   2137: '600-TX-433 APT O2 MONITOR - LOW LOW', class Tank Control Warnings, trigger "2062_Warning_Data_BTCS_WARNING_WORD_01" bit 9
   2138: 'TIT-436 2 PORT BWT TEMP - HIGH', class Tank Control Warnings, trigger "2062_Warning_Data_BTCS_WARNING_WORD_01" bit 10
   2139: 'TIT-436 2 STARBOARD BWT TEMP - HIGH', class Tank Control Warnings, trigger "2062_Warning_Data_BTCS_WARNING_WORD_01" bit 11
   2140: 'BTCS_WARNING_WORD_01_BIT_4', class Tank Control Warnings, trigger "2062_Warning_Data_BTCS_WARNING_WORD_01" bit 12
   2141: 'BTCS_WARNING_WORD_01_BIT_5', class Tank Control Warnings, trigger "2062_Warning_Data_BTCS_WARNING_WORD_01" bit 13
   2142: 'BTCS_WARNING_WORD_01_BIT_6', class Tank Control Warnings, trigger "2062_Warning_Data_BTCS_WARNING_WORD_01" bit 14
   2143: 'BTCS_WARNING_WORD_01_BIT_7', class Tank Control Warnings, trigger "2062_Warning_Data_BTCS_WARNING_WORD_01" bit 15
   2144: 'TT-426 1 FOR PEACK TANK TEMPERATURE - HIGH', class Tank Control Warnings, trigger "2062_Warning_Data_BTCS_WARNING_WORD_02" bit 0
   2145: 'TT-426 1 PORT TANK TEMPERATURE - HIGH', class Tank Control Warnings, trigger "2062_Warning_Data_BTCS_WARNING_WORD_02" bit 1
   2146: 'TT-426 1 STARBOARD TANK TEMPERATURE - HIGH', class Tank Control Warnings, trigger "2062_Warning_Data_BTCS_WARNING_WORD_02" bit 2
   2147: 'TT-426 3 PORT TANK TEMPERATURE - HIGH', class Tank Control Warnings, trigger "2062_Warning_Data_BTCS_WARNING_WORD_02" bit 3
   2148: 'TT-426 3 STARBOARD TANK TEMPERATURE - HIGH', class Tank Control Warnings, trigger "2062_Warning_Data_BTCS_WARNING_WORD_02" bit 4
   2149: 'TT-426 4 PORT TANK TEMPERATURE - HIGH', class Tank Control Warnings, trigger "2062_Warning_Data_BTCS_WARNING_WORD_02" bit 5
   2150: 'TT-426 4 STARBOARD TANK TEMPERATURE - HIGH', class Tank Control Warnings, trigger "2062_Warning_Data_BTCS_WARNING_WORD_02" bit 6
   2151: 'TT-426 5 PORT TANK TEMPERATURE - HIGH', class Tank Control Warnings, trigger "2062_Warning_Data_BTCS_WARNING_WORD_02" bit 7
   2152: 'PIT-415 2 PORT DECK IG PRESSURE - LOW', class Tank Control Warnings, trigger "2062_Warning_Data_BTCS_WARNING_WORD_02" bit 8
   2153: 'PIT-415 2 PORT DECK IG PRESSURE - HIGH', class Tank Control Warnings, trigger "2062_Warning_Data_BTCS_WARNING_WORD_02" bit 9
   2154: 'PIT-415 2 STARBOARD DECK IG PRESSURE - LOW', class Tank Control Warnings, trigger "2062_Warning_Data_BTCS_WARNING_WORD_02" bit 10
   2155: 'PIT-415 STARBOARD DECK IG PRESSURE - HIGH', class Tank Control Warnings, trigger "2062_Warning_Data_BTCS_WARNING_WORD_02" bit 11
   2156: 'PIT-424 2 PORT TANK PRESSURE - LOW', class Tank Control Warnings, trigger "2062_Warning_Data_BTCS_WARNING_WORD_02" bit 12
   2157: 'PIT-424 2 PORT TANK PRESSURE - HIGH', class Tank Control Warnings, trigger "2062_Warning_Data_BTCS_WARNING_WORD_02" bit 13
   2158: 'PIT-424 2 STARBOARD TANK PRESSURE - LOW', class Tank Control Warnings, trigger "2062_Warning_Data_BTCS_WARNING_WORD_02" bit 14
   2159: 'PIT-424 2 STARBOARD TANK PRESSURE - HIGH', class Tank Control Warnings, trigger "2062_Warning_Data_BTCS_WARNING_WORD_02" bit 15
   2160: 'FIT418 1 FOR PEACK TANK USD FLOW LOW', class Tank Control Warnings, trigger "2062_Warning_Data_BTCS_WARNING_WORD_03" bit 0
   2161: 'FIT418 1 FOR PEACK TANK USD FLOW HIGH', class Tank Control Warnings, trigger "2062_Warning_Data_BTCS_WARNING_WORD_03" bit 1
   2162: 'FIT418 1 PORT TANK USD FLOW LOW', class Tank Control Warnings, trigger "2062_Warning_Data_BTCS_WARNING_WORD_03" bit 2
   2163: 'FIT418 1 PORT TANK USD FLOW HIGH', class Tank Control Warnings, trigger "2062_Warning_Data_BTCS_WARNING_WORD_03" bit 3
   2164: 'FIT417 1 STARBOARD TANK USD FLOW LOW', class Tank Control Warnings, trigger "2062_Warning_Data_BTCS_WARNING_WORD_03" bit 4
   2165: 'FIT417 1 STARBOARD TANK USD FLOW HIGH', class Tank Control Warnings, trigger "2062_Warning_Data_BTCS_WARNING_WORD_03" bit 5
   2166: 'FIT418 3 PORT TANK USD FLOW LOW', class Tank Control Warnings, trigger "2062_Warning_Data_BTCS_WARNING_WORD_03" bit 6
   2167: 'FIT418 3 PORT TANK USD FLOW HIGH', class Tank Control Warnings, trigger "2062_Warning_Data_BTCS_WARNING_WORD_03" bit 7
   2168: 'TT-426 5 STARBOARD TANK TEMPERATURE - HIGH', class Tank Control Warnings, trigger "2062_Warning_Data_BTCS_WARNING_WORD_03" bit 8
   2169: 'TT-426 6 PORT TANK TEMPERATURE - HIGH', class Tank Control Warnings, trigger "2062_Warning_Data_BTCS_WARNING_WORD_03" bit 9
   2170: 'TT-426 6 STARBOARD TANK TEMPERATURE - HIGH', class Tank Control Warnings, trigger "2062_Warning_Data_BTCS_WARNING_WORD_03" bit 10
   2171: 'TT-426 7 AFT PEACK TANK TEMPERATURE - HIGH', class Tank Control Warnings, trigger "2062_Warning_Data_BTCS_WARNING_WORD_03" bit 11
   2172: 'BTCS_WARNING_WORD_03_BIT_4', class Tank Control Warnings, trigger "2062_Warning_Data_BTCS_WARNING_WORD_03" bit 12
   2173: 'BTCS_WARNING_WORD_03_BIT_5', class Tank Control Warnings, trigger "2062_Warning_Data_BTCS_WARNING_WORD_03" bit 13
   2174: 'BTCS_WARNING_WORD_03_BIT_6', class Tank Control Warnings, trigger "2062_Warning_Data_BTCS_WARNING_WORD_03" bit 14
   2175: 'BTCS_WARNING_WORD_03_BIT_7', class Tank Control Warnings, trigger "2062_Warning_Data_BTCS_WARNING_WORD_03" bit 15
   2176: 'FIT417 5 STARBOARD TANK USD FLOW LOW', class Tank Control Warnings, trigger "2062_Warning_Data_BTCS_WARNING_WORD_04" bit 0
   2177: 'FIT417 5 STARBOARD TANK USD FLOW HIGH', class Tank Control Warnings, trigger "2062_Warning_Data_BTCS_WARNING_WORD_04" bit 1
   2178: 'FIT418 6 PORT TANK USD FLOW LOW', class Tank Control Warnings, trigger "2062_Warning_Data_BTCS_WARNING_WORD_04" bit 2
   2179: 'FIT418 6 PORT TANK USD FLOW HIGH', class Tank Control Warnings, trigger "2062_Warning_Data_BTCS_WARNING_WORD_04" bit 3
   2180: 'FIT417 6 STARBOARD TANK USD FLOW LOW', class Tank Control Warnings, trigger "2062_Warning_Data_BTCS_WARNING_WORD_04" bit 4
   2181: 'FIT417 6 STARBOARD TANK USD FLOW HIGH', class Tank Control Warnings, trigger "2062_Warning_Data_BTCS_WARNING_WORD_04" bit 5
   2182: 'FIT418 7 APT TANK USD FLOW LOW', class Tank Control Warnings, trigger "2062_Warning_Data_BTCS_WARNING_WORD_04" bit 6
   2183: 'FIT418 7 APT TANK USD FLOW HIGH', class Tank Control Warnings, trigger "2062_Warning_Data_BTCS_WARNING_WORD_04" bit 7
   2184: 'FIT417 3 STARBOARD TANK USD FLOW LOW', class Tank Control Warnings, trigger "2062_Warning_Data_BTCS_WARNING_WORD_04" bit 8
   2185: 'FIT417 3 STARBOARD TANK USD FLOW HIGH', class Tank Control Warnings, trigger "2062_Warning_Data_BTCS_WARNING_WORD_04" bit 9
   2186: 'FIT418 4 PORT TANK USD FLOW LOW', class Tank Control Warnings, trigger "2062_Warning_Data_BTCS_WARNING_WORD_04" bit 10
   2187: 'FIT418 4 PORT TANK USD FLOW HIGH', class Tank Control Warnings, trigger "2062_Warning_Data_BTCS_WARNING_WORD_04" bit 11
   2188: 'FIT417 4 STARBOARD TANK USD FLOW LOW', class Tank Control Warnings, trigger "2062_Warning_Data_BTCS_WARNING_WORD_04" bit 12
   2189: 'FIT417 4 STARBOARD TANK USD FLOW HIGH', class Tank Control Warnings, trigger "2062_Warning_Data_BTCS_WARNING_WORD_04" bit 13
   2190: 'FIT418 5 PORT TANK USD FLOW LOW', class Tank Control Warnings, trigger "2062_Warning_Data_BTCS_WARNING_WORD_04" bit 14
   2191: 'FIT418 5 PORT TANK USD FLOW HIGH', class Tank Control Warnings, trigger "2062_Warning_Data_BTCS_WARNING_WORD_04" bit 15
   2192: 'FIT419 3 STARBOARD MBG FLOW LOW', class Tank Control Warnings, trigger "2062_Warning_Data_BTCS_WARNING_WORD_05" bit 0
   2193: 'FIT419 3 STARBOARD MBG FLOW HIGH', class Tank Control Warnings, trigger "2062_Warning_Data_BTCS_WARNING_WORD_05" bit 1
   2194: 'FIT420 4 PORT MBG FLOW LOW', class Tank Control Warnings, trigger "2062_Warning_Data_BTCS_WARNING_WORD_05" bit 2
   2195: 'FIT420 4 PORT MBG FLOW HIGH', class Tank Control Warnings, trigger "2062_Warning_Data_BTCS_WARNING_WORD_05" bit 3
   2196: 'FIT419 4 STARBOARD MBG FLOW LOW', class Tank Control Warnings, trigger "2062_Warning_Data_BTCS_WARNING_WORD_05" bit 4
   2197: 'FIT419 4 STARBOARD MBG FLOW HIGH', class Tank Control Warnings, trigger "2062_Warning_Data_BTCS_WARNING_WORD_05" bit 5
   2198: 'FIT420 5 PORT MBG FLOW LOW', class Tank Control Warnings, trigger "2062_Warning_Data_BTCS_WARNING_WORD_05" bit 6
   2199: 'FIT420 5 PORT MBG FLOW HIGH', class Tank Control Warnings, trigger "2062_Warning_Data_BTCS_WARNING_WORD_05" bit 7
   2200: 'FIT420 1 FPT MBG FLOW LOW', class Tank Control Warnings, trigger "2062_Warning_Data_BTCS_WARNING_WORD_05" bit 8
   2201: 'FIT420 1 FPT MBG FLOW HIGH', class Tank Control Warnings, trigger "2062_Warning_Data_BTCS_WARNING_WORD_05" bit 9
   2202: 'FIT420 1 PORT MBG FLOW LOW', class Tank Control Warnings, trigger "2062_Warning_Data_BTCS_WARNING_WORD_05" bit 10
   2203: 'FIT420 1 PORT MBG FLOW HIGH', class Tank Control Warnings, trigger "2062_Warning_Data_BTCS_WARNING_WORD_05" bit 11
   2204: 'FIT419 1 STARBOARD MBG FLOW LOW', class Tank Control Warnings, trigger "2062_Warning_Data_BTCS_WARNING_WORD_05" bit 12
   2205: 'FIT419 1 STARBOARD MBG FLOW HIGH', class Tank Control Warnings, trigger "2062_Warning_Data_BTCS_WARNING_WORD_05" bit 13
   2206: 'FIT420 3 PORT MBG FLOW LOW', class Tank Control Warnings, trigger "2062_Warning_Data_BTCS_WARNING_WORD_05" bit 14
   2207: 'FIT420 3 PORT MBG FLOW HIGH', class Tank Control Warnings, trigger "2062_Warning_Data_BTCS_WARNING_WORD_05" bit 15
   2208: 'PT415 RIO1 DECK IG PRESSURE LOW', class Tank Control Warnings, trigger "2062_Warning_Data_BTCS_WARNING_WORD_06" bit 0
   2209: 'PT415 RIO1 DECK IG PRESSURE HIGH', class Tank Control Warnings, trigger "2062_Warning_Data_BTCS_WARNING_WORD_06" bit 1
   2210: 'PT415 RIO3 DECK IG PRESSURE LOW', class Tank Control Warnings, trigger "2062_Warning_Data_BTCS_WARNING_WORD_06" bit 2
   2211: 'PT415 RIO3 DECK IG PRESSURE HIGH', class Tank Control Warnings, trigger "2062_Warning_Data_BTCS_WARNING_WORD_06" bit 3
   2212: 'PT415 RIO4 DECK IG PRESSURE LOW', class Tank Control Warnings, trigger "2062_Warning_Data_BTCS_WARNING_WORD_06" bit 4
   2213: 'PT415 RIO4 DECK IG PRESSURE HIGH', class Tank Control Warnings, trigger "2062_Warning_Data_BTCS_WARNING_WORD_06" bit 5
   2214: 'PT415 RIO5 DECK IG PRESSURE LOW', class Tank Control Warnings, trigger "2062_Warning_Data_BTCS_WARNING_WORD_06" bit 6
   2215: 'PT415 RIO5 DECK IG PRESSURE HIGH', class Tank Control Warnings, trigger "2062_Warning_Data_BTCS_WARNING_WORD_06" bit 7
   2216: 'FIT419 5 STARBOARD MBG FLOW LOW', class Tank Control Warnings, trigger "2062_Warning_Data_BTCS_WARNING_WORD_06" bit 8
   2217: 'FIT419 5 STARBOARD MBG FLOW HIGH', class Tank Control Warnings, trigger "2062_Warning_Data_BTCS_WARNING_WORD_06" bit 9
   2218: 'FIT420 6 PORT MBG FLOW LOW', class Tank Control Warnings, trigger "2062_Warning_Data_BTCS_WARNING_WORD_06" bit 10
   2219: 'FIT420 6 PORT MBG FLOW HIGH', class Tank Control Warnings, trigger "2062_Warning_Data_BTCS_WARNING_WORD_06" bit 11
   2220: 'FIT419 6 STARBOARD MBG FLOW LOW', class Tank Control Warnings, trigger "2062_Warning_Data_BTCS_WARNING_WORD_06" bit 12
   2221: 'FIT419 6 STARBOARD MBG FLOW HIGH', class Tank Control Warnings, trigger "2062_Warning_Data_BTCS_WARNING_WORD_06" bit 13
   2222: 'FIT420 7 APT MBG FLOW LOW', class Tank Control Warnings, trigger "2062_Warning_Data_BTCS_WARNING_WORD_06" bit 14
   2223: 'FIT420 7 APT MBG FLOW HIGH', class Tank Control Warnings, trigger "2062_Warning_Data_BTCS_WARNING_WORD_06" bit 15
   2224: 'PIT424 RIO5 TANK PRESSURE LOW', class Tank Control Warnings, trigger "2062_Warning_Data_BTCS_WARNING_WORD_07" bit 0
   2225: 'PIT424 RIO5 TANK PRESSURE HIGH', class Tank Control Warnings, trigger "2062_Warning_Data_BTCS_WARNING_WORD_07" bit 1
   2226: 'PIT424 RIO6 TANK PRESSURE LOW', class Tank Control Warnings, trigger "2062_Warning_Data_BTCS_WARNING_WORD_07" bit 2
   2227: 'PIT424 RIO6 TANK PRESSURE HIGH', class Tank Control Warnings, trigger "2062_Warning_Data_BTCS_WARNING_WORD_07" bit 3
   2228: 'PIT424 RIO7 TANK PRESSURE LOW', class Tank Control Warnings, trigger "2062_Warning_Data_BTCS_WARNING_WORD_07" bit 4
   2229: 'PIT424 RIO7 TANK PRESSURE HIGH', class Tank Control Warnings, trigger "2062_Warning_Data_BTCS_WARNING_WORD_07" bit 5
   2230: 'BTCS_WARNING_WORD_07_BIT_14', class Tank Control Warnings, trigger "2062_Warning_Data_BTCS_WARNING_WORD_07" bit 6
   2231: 'BTCS_WARNING_WORD_07_BIT_15', class Tank Control Warnings, trigger "2062_Warning_Data_BTCS_WARNING_WORD_07" bit 7
   2232: 'PT415 RIO6 DECK IG PRESSURE LOW', class Tank Control Warnings, trigger "2062_Warning_Data_BTCS_WARNING_WORD_07" bit 8
   2233: 'PT415 RIO6 DECK IG PRESSURE HIGH', class Tank Control Warnings, trigger "2062_Warning_Data_BTCS_WARNING_WORD_07" bit 9
   2234: 'PIT424 RIO1 TANK PRESSURE LOW', class Tank Control Warnings, trigger "2062_Warning_Data_BTCS_WARNING_WORD_07" bit 10
   2235: 'PIT424 RIO1 TANK PRESSURE HIGH', class Tank Control Warnings, trigger "2062_Warning_Data_BTCS_WARNING_WORD_07" bit 11
   2236: 'PIT424 RIO3 TANK PRESSURE LOW', class Tank Control Warnings, trigger "2062_Warning_Data_BTCS_WARNING_WORD_07" bit 12
   2237: 'PIT424 RIO3 TANK PRESSURE HIGH', class Tank Control Warnings, trigger "2062_Warning_Data_BTCS_WARNING_WORD_07" bit 13
   2238: 'PIT424 RIO4 TANK PRESSURE LOW', class Tank Control Warnings, trigger "2062_Warning_Data_BTCS_WARNING_WORD_07" bit 14
   2239: 'PIT424 RIO4 TANK PRESSURE HIGH', class Tank Control Warnings, trigger "2062_Warning_Data_BTCS_WARNING_WORD_07" bit 15
   2240: 'LS425 4 STARBOARD TANK LEVEL HIGH HIGH', class Tank Control Warnings, trigger "2062_Warning_Data_BTCS_WARNING_WORD_08" bit 0
   2241: 'LS425 5 PORT TANK LEVEL HIGH HIGH', class Tank Control Warnings, trigger "2062_Warning_Data_BTCS_WARNING_WORD_08" bit 1
   2242: 'LS425 5 STARBOARD TANK LEVEL HIGH HIGH', class Tank Control Warnings, trigger "2062_Warning_Data_BTCS_WARNING_WORD_08" bit 2
   2243: 'LS425 6 PORT TANK LEVEL HIGH HIGH', class Tank Control Warnings, trigger "2062_Warning_Data_BTCS_WARNING_WORD_08" bit 3
   2244: 'LS425 6 STARBOARD TANK LEVEL HIGH HIGH', class Tank Control Warnings, trigger "2062_Warning_Data_BTCS_WARNING_WORD_08" bit 4
   2245: 'LS425 AP TANK LEVEL HIGH HIGH', class Tank Control Warnings, trigger "2062_Warning_Data_BTCS_WARNING_WORD_08" bit 5
   2246: 'BTCS_WARNING_WORD_08_BIT_14', class Tank Control Warnings, trigger "2062_Warning_Data_BTCS_WARNING_WORD_08" bit 6
   2247: 'LS425 FP TANK LEVEL HIGH HIGH', class Tank Control Warnings, trigger "2062_Warning_Data_BTCS_WARNING_WORD_08" bit 7
   2248: 'PT415 RIO7 DECK IG PRESSURE LOW', class Tank Control Warnings, trigger "2062_Warning_Data_BTCS_WARNING_WORD_08" bit 8
   2249: 'PT415 RIO7 DECK IG PRESSURE HIGH', class Tank Control Warnings, trigger "2062_Warning_Data_BTCS_WARNING_WORD_08" bit 9
   2250: 'LS425 1 STARBOARD TANK LEVEL HIGH HIGH', class Tank Control Warnings, trigger "2062_Warning_Data_BTCS_WARNING_WORD_08" bit 10
   2251: 'LS425 2 PORT TANK LEVEL HIGH HIGH', class Tank Control Warnings, trigger "2062_Warning_Data_BTCS_WARNING_WORD_08" bit 11
   2252: 'LS425 2 STARBOARD TANK LEVEL HIGH HIGH', class Tank Control Warnings, trigger "2062_Warning_Data_BTCS_WARNING_WORD_08" bit 12
   2253: 'LS425 3 PORT TANK LEVEL HIGH HIGH', class Tank Control Warnings, trigger "2062_Warning_Data_BTCS_WARNING_WORD_08" bit 13
   2254: 'LS425 3 STARBOARD TANK LEVEL HIGH HIGH', class Tank Control Warnings, trigger "2062_Warning_Data_BTCS_WARNING_WORD_08" bit 14
   2255: 'LS425 4 PORT TANK LEVEL HIGH HIGH', class Tank Control Warnings, trigger "2062_Warning_Data_BTCS_WARNING_WORD_08" bit 15
   2256: 'LT422 FPT TANK LEVEL HIGH', class Tank Control Warnings, trigger "2062_Warning_Data_BTCS_WARNING_WORD_09" bit 0
   2257: 'LT422 FPT TANK LEVEL LOW', class Tank Control Warnings, trigger "2062_Warning_Data_BTCS_WARNING_WORD_09" bit 1
   2258: 'LT422 1 PORT TANK LEVEL HIGH', class Tank Control Warnings, trigger "2062_Warning_Data_BTCS_WARNING_WORD_09" bit 2
   2259: 'LT422 1 PORT TANK LEVEL LOW', class Tank Control Warnings, trigger "2062_Warning_Data_BTCS_WARNING_WORD_09" bit 3
   2260: 'LT422 1 STARBOARD TANK LEVEL HIGH', class Tank Control Warnings, trigger "2062_Warning_Data_BTCS_WARNING_WORD_09" bit 4
   2261: 'LT422 1 STARBOARD TANK LEVEL LOW', class Tank Control Warnings, trigger "2062_Warning_Data_BTCS_WARNING_WORD_09" bit 5
   2262: 'LT422 2 PORT TANK LEVEL HIGH', class Tank Control Warnings, trigger "2062_Warning_Data_BTCS_WARNING_WORD_09" bit 6
   2263: 'LT422 2 PORT TANK LEVEL LOW', class Tank Control Warnings, trigger "2062_Warning_Data_BTCS_WARNING_WORD_09" bit 7
   2264: 'PS436 RIO1 TANK GROUP PRESURE HIGH HIGH', class Tank Control Warnings, trigger "2062_Warning_Data_BTCS_WARNING_WORD_09" bit 8
   2265: 'PS436 RIO2 TANK GROUP PRESURE HIGH HIGH', class Tank Control Warnings, trigger "2062_Warning_Data_BTCS_WARNING_WORD_09" bit 9
   2266: 'PS436 RIO3 TANK GROUP PRESURE HIGH HIGH', class Tank Control Warnings, trigger "2062_Warning_Data_BTCS_WARNING_WORD_09" bit 10
   2267: 'PS436 RIO4 TANK GROUP PRESURE HIGH HIGH', class Tank Control Warnings, trigger "2062_Warning_Data_BTCS_WARNING_WORD_09" bit 11
   2268: 'PS436 RIO5 TANK GROUP PRESURE HIGH HIGH', class Tank Control Warnings, trigger "2062_Warning_Data_BTCS_WARNING_WORD_09" bit 12
   2269: 'PS436 RIO6 TANK GROUP PRESURE HIGH HIGH', class Tank Control Warnings, trigger "2062_Warning_Data_BTCS_WARNING_WORD_09" bit 13
   2270: 'PS436 RIO7 TANK GROUP PRESURE HIGH HIGH', class Tank Control Warnings, trigger "2062_Warning_Data_BTCS_WARNING_WORD_09" bit 14
   2271: 'LS425 1 PORT TANK LEVEL HIGH HIGH', class Tank Control Warnings, trigger "2062_Warning_Data_BTCS_WARNING_WORD_09" bit 15
   2272: 'LT422 4 STARBOARD TANK LEVEL HIGH', class Tank Control Warnings, trigger "2062_Warning_Data_BTCS_WARNING_WORD_10" bit 0
   2273: 'LT422 4 STARBOARD TANK LEVEL LOW', class Tank Control Warnings, trigger "2062_Warning_Data_BTCS_WARNING_WORD_10" bit 1
   2274: 'LT422 5 PORT TANK LEVEL HIGH', class Tank Control Warnings, trigger "2062_Warning_Data_BTCS_WARNING_WORD_10" bit 2
   2275: 'LT422 5 PORT TANK LEVEL LOW', class Tank Control Warnings, trigger "2062_Warning_Data_BTCS_WARNING_WORD_10" bit 3
   2276: 'LT422 5 STARBOARD TANK LEVEL HIGH', class Tank Control Warnings, trigger "2062_Warning_Data_BTCS_WARNING_WORD_10" bit 4
   2277: 'LT422 5 STARBOARD TANK LEVEL LOW', class Tank Control Warnings, trigger "2062_Warning_Data_BTCS_WARNING_WORD_10" bit 5
   2278: 'LT422 6 PORT TANK LEVEL HIGH', class Tank Control Warnings, trigger "2062_Warning_Data_BTCS_WARNING_WORD_10" bit 6
   2279: 'LT422 6 PORT TANK LEVEL LOW', class Tank Control Warnings, trigger "2062_Warning_Data_BTCS_WARNING_WORD_10" bit 7
   2280: 'LT422 2 STARBOARD TANK LEVEL HIGH', class Tank Control Warnings, trigger "2062_Warning_Data_BTCS_WARNING_WORD_10" bit 8
   2281: 'LT422 2 STARBOARD TANK LEVEL LOW', class Tank Control Warnings, trigger "2062_Warning_Data_BTCS_WARNING_WORD_10" bit 9
   2282: 'LT422 3 PORT TANK LEVEL HIGH', class Tank Control Warnings, trigger "2062_Warning_Data_BTCS_WARNING_WORD_10" bit 10
   2283: 'LT422 3 PORT TANK LEVEL LOW', class Tank Control Warnings, trigger "2062_Warning_Data_BTCS_WARNING_WORD_10" bit 11
   2284: 'LT422 3 STARBOARD TANK LEVEL HIGH', class Tank Control Warnings, trigger "2062_Warning_Data_BTCS_WARNING_WORD_10" bit 12
   2285: 'LT422 3 STARBOARD TANK LEVEL LOW', class Tank Control Warnings, trigger "2062_Warning_Data_BTCS_WARNING_WORD_10" bit 13
   2286: 'LT422 4 PORT TANK LEVEL HIGH', class Tank Control Warnings, trigger "2062_Warning_Data_BTCS_WARNING_WORD_10" bit 14
   2287: 'LT422 4 PORT TANK LEVEL LOW', class Tank Control Warnings, trigger "2062_Warning_Data_BTCS_WARNING_WORD_10" bit 15
   2288: 'TT426 2S BWT TEMP HIGH', class Tank Control Warnings, trigger "2062_Warning_Data_BTCS_WARNING_WORD_11" bit 0
   2289: 'TT426 3P BWT TEMP HIGH', class Tank Control Warnings, trigger "2062_Warning_Data_BTCS_WARNING_WORD_11" bit 1
   2290: 'TT426 3S BWT TEMP HIGH', class Tank Control Warnings, trigger "2062_Warning_Data_BTCS_WARNING_WORD_11" bit 2
   2291: 'TT426 4P BWT TEMP HIGH', class Tank Control Warnings, trigger "2062_Warning_Data_BTCS_WARNING_WORD_11" bit 3
   2292: 'TT426 4S BWT TEMP HIGH', class Tank Control Warnings, trigger "2062_Warning_Data_BTCS_WARNING_WORD_11" bit 4
   2293: 'TT426 5P BWT TEMP HIGH', class Tank Control Warnings, trigger "2062_Warning_Data_BTCS_WARNING_WORD_11" bit 5
   2294: 'TT426 5S BWT TEMP HIGH', class Tank Control Warnings, trigger "2062_Warning_Data_BTCS_WARNING_WORD_11" bit 6
   2295: 'TT426 6P BWT TEMP HIGH', class Tank Control Warnings, trigger "2062_Warning_Data_BTCS_WARNING_WORD_11" bit 7
   2296: 'LT422 6S TANK LEVEL HIGH', class Tank Control Warnings, trigger "2062_Warning_Data_BTCS_WARNING_WORD_11" bit 8
   2297: 'LT422 6S TANK LEVEL LOW', class Tank Control Warnings, trigger "2062_Warning_Data_BTCS_WARNING_WORD_11" bit 9
   2298: 'LT422 APT TANK LEVEL HIGH', class Tank Control Warnings, trigger "2062_Warning_Data_BTCS_WARNING_WORD_11" bit 10
   2299: 'LT422 APT TANK LEVEL LOW', class Tank Control Warnings, trigger "2062_Warning_Data_BTCS_WARNING_WORD_11" bit 11
   2300: 'TT426 FPT BWT TEMP HIGH', class Tank Control Warnings, trigger "2062_Warning_Data_BTCS_WARNING_WORD_11" bit 12
   2301: 'TT426 1P BWT TEMP HIGH', class Tank Control Warnings, trigger "2062_Warning_Data_BTCS_WARNING_WORD_11" bit 13
   2302: 'TT426 1S BWT TEMP HIGH', class Tank Control Warnings, trigger "2062_Warning_Data_BTCS_WARNING_WORD_11" bit 14
   2303: 'TT426 2P BWT TEMP HIGH', class Tank Control Warnings, trigger "2062_Warning_Data_BTCS_WARNING_WORD_11" bit 15
   2304: 'FIT417 3S USD OUT OF RANGE', class Tank Control Warnings, trigger "2062_Warning_Data_BTCS_WARNING_WORD_12" bit 0
   2305: 'FIT418 4P USD OUT OF RANGE', class Tank Control Warnings, trigger "2062_Warning_Data_BTCS_WARNING_WORD_12" bit 1
   2306: 'FIT417 4S USD OUT OF RANGE', class Tank Control Warnings, trigger "2062_Warning_Data_BTCS_WARNING_WORD_12" bit 2
   2307: 'FIT418 5P USD OUT OF RANGE', class Tank Control Warnings, trigger "2062_Warning_Data_BTCS_WARNING_WORD_12" bit 3
   2308: 'FIT417 5S USD OUT OF RANGE', class Tank Control Warnings, trigger "2062_Warning_Data_BTCS_WARNING_WORD_12" bit 4
   2309: 'FIT418 6P USD OUT OF RANGE', class Tank Control Warnings, trigger "2062_Warning_Data_BTCS_WARNING_WORD_12" bit 5
   2310: 'FIT417 6S USD OUT OF RANGE', class Tank Control Warnings, trigger "2062_Warning_Data_BTCS_WARNING_WORD_12" bit 6
   2311: 'FIT417 APT USD OUT OF RANGE', class Tank Control Warnings, trigger "2062_Warning_Data_BTCS_WARNING_WORD_12" bit 7
   2312: 'TT426 6S BWT TEMP OUT OF RANGE', class Tank Control Warnings, trigger "2062_Warning_Data_BTCS_WARNING_WORD_12" bit 8
   2313: 'TT426 APT BWT TEMP OUT OF RANGE', class Tank Control Warnings, trigger "2062_Warning_Data_BTCS_WARNING_WORD_12" bit 9
   2314: 'FIT418 FPT USD OUT OF RANGE', class Tank Control Warnings, trigger "2062_Warning_Data_BTCS_WARNING_WORD_12" bit 10
   2315: 'FIT418 1P USD OUT OF RANGE', class Tank Control Warnings, trigger "2062_Warning_Data_BTCS_WARNING_WORD_12" bit 11
   2316: 'FIT417 1S USD OUT OF RANGE', class Tank Control Warnings, trigger "2062_Warning_Data_BTCS_WARNING_WORD_12" bit 12
   2317: 'FIT418 2P USD OUT OF RANGE', class Tank Control Warnings, trigger "2062_Warning_Data_BTCS_WARNING_WORD_12" bit 13
   2318: 'FIT417 2S USD OUT OF RANGE', class Tank Control Warnings, trigger "2062_Warning_Data_BTCS_WARNING_WORD_12" bit 14
   2319: 'FIT418 3P USD OUT OF RANGE', class Tank Control Warnings, trigger "2062_Warning_Data_BTCS_WARNING_WORD_12" bit 15
   2320: 'FIT419 4S MBG FLOW OUT OF RANGE', class Tank Control Warnings, trigger "2062_Warning_Data_BTCS_WARNING_WORD_13" bit 0
   2321: 'FIT420 5P MBG FLOW OUT OF RANGE', class Tank Control Warnings, trigger "2062_Warning_Data_BTCS_WARNING_WORD_13" bit 1
   2322: 'FIT419 5S MBG FLOW OUT OF RANGE', class Tank Control Warnings, trigger "2062_Warning_Data_BTCS_WARNING_WORD_13" bit 2
   2323: 'FIT420 6P MBG FLOW OUT OF RANGE', class Tank Control Warnings, trigger "2062_Warning_Data_BTCS_WARNING_WORD_13" bit 3
   2324: 'FIT419 6S MBG FLOW OUT OF RANGE', class Tank Control Warnings, trigger "2062_Warning_Data_BTCS_WARNING_WORD_13" bit 4
   2325: 'FIT420 APT MBG FLOW OUT OF RANGE', class Tank Control Warnings, trigger "2062_Warning_Data_BTCS_WARNING_WORD_13" bit 5
   2326: 'PT415 RIO1 DECK IG PRESSURE OUT OF RANGE', class Tank Control Warnings, trigger "2062_Warning_Data_BTCS_WARNING_WORD_13" bit 6
   2327: 'PT415 RIO2 DECK IG PRESSURE OUT OF RANGE', class Tank Control Warnings, trigger "2062_Warning_Data_BTCS_WARNING_WORD_13" bit 7
   2328: 'FIT420 FPT MBG FLOW OUT OF RANGE', class Tank Control Warnings, trigger "2062_Warning_Data_BTCS_WARNING_WORD_13" bit 8
   2329: 'FIT420 1P MBG FLOW OUT OF RANGE', class Tank Control Warnings, trigger "2062_Warning_Data_BTCS_WARNING_WORD_13" bit 9
   2330: 'FIT419 1S MBG FLOW OUT OF RANGE', class Tank Control Warnings, trigger "2062_Warning_Data_BTCS_WARNING_WORD_13" bit 10
   2331: 'FIT420 2P MBG FLOW OUT OF RANGE', class Tank Control Warnings, trigger "2062_Warning_Data_BTCS_WARNING_WORD_13" bit 11
   2332: 'FIT419 2S MBG FLOW OUT OF RANGE', class Tank Control Warnings, trigger "2062_Warning_Data_BTCS_WARNING_WORD_13" bit 12
   2333: 'FIT420 3P MBG FLOW OUT OF RANGE', class Tank Control Warnings, trigger "2062_Warning_Data_BTCS_WARNING_WORD_13" bit 13
   2334: 'FIT419 3S MBG FLOW OUT OF RANGE', class Tank Control Warnings, trigger "2062_Warning_Data_BTCS_WARNING_WORD_13" bit 14
   2335: 'FIT420 4P MBG FLOW OUT OF RANGE', class Tank Control Warnings, trigger "2062_Warning_Data_BTCS_WARNING_WORD_13" bit 15
   2336: 'PIT424 RIO4 TANK PRESSURE OUT OF RANGE', class Tank Control Warnings, trigger "2062_Warning_Data_BTCS_WARNING_WORD_14" bit 0
   2337: 'PIT424 RIO5 TANK PRESSURE OUT OF RANGE', class Tank Control Warnings, trigger "2062_Warning_Data_BTCS_WARNING_WORD_14" bit 1
   2338: 'PIT424 RIO6 TANK PRESSURE OUT OF RANGE', class Tank Control Warnings, trigger "2062_Warning_Data_BTCS_WARNING_WORD_14" bit 2
   2339: 'PIT424 RIO7 TANK PRESSURE OUT OF RANGE', class Tank Control Warnings, trigger "2062_Warning_Data_BTCS_WARNING_WORD_14" bit 3
   2340: 'LT422 FPT TANK LEVEL OUT OF RANGE', class Tank Control Warnings, trigger "2062_Warning_Data_BTCS_WARNING_WORD_14" bit 4
   2341: 'LT422 1P TANK LEVEL OUT OF RANGE', class Tank Control Warnings, trigger "2062_Warning_Data_BTCS_WARNING_WORD_14" bit 5
   2342: 'LT422 1S TANK LEVEL OUT OF RANGE', class Tank Control Warnings, trigger "2062_Warning_Data_BTCS_WARNING_WORD_14" bit 6
   2343: 'LT422 2P TANK LEVEL OUT OF RANGE', class Tank Control Warnings, trigger "2062_Warning_Data_BTCS_WARNING_WORD_14" bit 7
   2344: 'PT415 RIO3 DECK IG PRESSURE OUT OF RANGE', class Tank Control Warnings, trigger "2062_Warning_Data_BTCS_WARNING_WORD_14" bit 8
   2345: 'PT415 RIO4 DECK IG PRESSURE OUT OF RANGE', class Tank Control Warnings, trigger "2062_Warning_Data_BTCS_WARNING_WORD_14" bit 9
   2346: 'PT415 RIO5 DECK IG PRESSURE OUT OF RANGE', class Tank Control Warnings, trigger "2062_Warning_Data_BTCS_WARNING_WORD_14" bit 10
   2347: 'PT415 RIO6 DECK IG PRESSURE OUT OF RANGE', class Tank Control Warnings, trigger "2062_Warning_Data_BTCS_WARNING_WORD_14" bit 11
   2348: 'PT415 RIO7 DECK IG PRESSURE OUT OF RANGE', class Tank Control Warnings, trigger "2062_Warning_Data_BTCS_WARNING_WORD_14" bit 12
   2349: 'PIT424 RIO1 TANK PRESSURE OUT OF RANGE', class Tank Control Warnings, trigger "2062_Warning_Data_BTCS_WARNING_WORD_14" bit 13
   2350: 'PIT424 RIO2 TANK PRESSURE OUT OF RANGE', class Tank Control Warnings, trigger "2062_Warning_Data_BTCS_WARNING_WORD_14" bit 14
   2351: 'PIT424 RIO3 TANK PRESSURE OUT OF RANGE', class Tank Control Warnings, trigger "2062_Warning_Data_BTCS_WARNING_WORD_14" bit 15
   2352: 'LT422 6S TANK LEVEL OUT OF RANGE', class Tank Control Warnings, trigger "2062_Warning_Data_BTCS_WARNING_WORD_15" bit 0
   2353: 'LT422 APT TANK LEVEL OUT OF RANGE', class Tank Control Warnings, trigger "2062_Warning_Data_BTCS_WARNING_WORD_15" bit 1
   2354: '600-TX-433 APT O2 MONITOR OUT OF RANGE', class Tank Control Warnings, trigger "2062_Warning_Data_BTCS_WARNING_WORD_15" bit 2
   2355: 'PH426 FPT OUT OF RANGE', class Tank Control Warnings, trigger "2062_Warning_Data_BTCS_WARNING_WORD_15" bit 3
   2356: 'PH426 1P OUT OF RANGE', class Tank Control Warnings, trigger "2062_Warning_Data_BTCS_WARNING_WORD_15" bit 4
   2357: 'PH426 1S OUT OF RANGE', class Tank Control Warnings, trigger "2062_Warning_Data_BTCS_WARNING_WORD_15" bit 5
   2358: 'PH426 2P OUT OF RANGE', class Tank Control Warnings, trigger "2062_Warning_Data_BTCS_WARNING_WORD_15" bit 6
   2359: 'PH426 2S OUT OF RANGE', class Tank Control Warnings, trigger "2062_Warning_Data_BTCS_WARNING_WORD_15" bit 7
   2360: 'LT422 2S TANK LEVEL OUT OF RANGE', class Tank Control Warnings, trigger "2062_Warning_Data_BTCS_WARNING_WORD_15" bit 8
   2361: 'LT422 3P TANK LEVEL OUT OF RANGE', class Tank Control Warnings, trigger "2062_Warning_Data_BTCS_WARNING_WORD_15" bit 9
   2362: 'LT422 3S TANK LEVEL OUT OF RANGE', class Tank Control Warnings, trigger "2062_Warning_Data_BTCS_WARNING_WORD_15" bit 10
   2363: 'LT422 4P TANK LEVEL OUT OF RANGE', class Tank Control Warnings, trigger "2062_Warning_Data_BTCS_WARNING_WORD_15" bit 11
   2364: 'LT422 4S TANK LEVEL OUT OF RANGE', class Tank Control Warnings, trigger "2062_Warning_Data_BTCS_WARNING_WORD_15" bit 12
   2365: 'LT422 5P TANK LEVEL OUT OF RANGE', class Tank Control Warnings, trigger "2062_Warning_Data_BTCS_WARNING_WORD_15" bit 13
   2366: 'LT422 5S TANK LEVEL OUT OF RANGE', class Tank Control Warnings, trigger "2062_Warning_Data_BTCS_WARNING_WORD_15" bit 14
   2367: 'LT422 6P TANK LEVEL OUT OF RANGE', class Tank Control Warnings, trigger "2062_Warning_Data_BTCS_WARNING_WORD_15" bit 15
   2368: 'PH425 6S OUT OF RANGE', class Tank Control Warnings, trigger "2062_Warning_Data_BTCS_WARNING_WORD_16" bit 0
   2369: 'PH426 APT OUT OF RANGE', class Tank Control Warnings, trigger "2062_Warning_Data_BTCS_WARNING_WORD_16" bit 1
   2370: 'DO428 FPT OUT OF RANGE', class Tank Control Warnings, trigger "2062_Warning_Data_BTCS_WARNING_WORD_16" bit 2
   2371: 'DO428 1P OUT OF RANGE', class Tank Control Warnings, trigger "2062_Warning_Data_BTCS_WARNING_WORD_16" bit 3
   2372: 'DO427 1S OUT OF RANGE', class Tank Control Warnings, trigger "2062_Warning_Data_BTCS_WARNING_WORD_16" bit 4
   2373: 'DO428 2P OUT OF RANGE', class Tank Control Warnings, trigger "2062_Warning_Data_BTCS_WARNING_WORD_16" bit 5
   2374: 'DO427 2S OUT OF RANGE', class Tank Control Warnings, trigger "2062_Warning_Data_BTCS_WARNING_WORD_16" bit 6
   2375: 'DO428 3P OUT OF RANGE', class Tank Control Warnings, trigger "2062_Warning_Data_BTCS_WARNING_WORD_16" bit 7
   2376: 'PH426 3P OUT OF RANGE', class Tank Control Warnings, trigger "2062_Warning_Data_BTCS_WARNING_WORD_16" bit 8
   2377: 'PH425 3S OUT OF RANGE', class Tank Control Warnings, trigger "2062_Warning_Data_BTCS_WARNING_WORD_16" bit 9
   2378: 'PH426 4P OUT OF RANGE', class Tank Control Warnings, trigger "2062_Warning_Data_BTCS_WARNING_WORD_16" bit 10
   2379: '', class Tank Control Warnings, trigger "2062_Warning_Data_BTCS_WARNING_WORD_16" bit 11
   2380: 'PH425 4S OUT OF RANGE', class Tank Control Warnings, trigger "2062_Warning_Data_BTCS_WARNING_WORD_16" bit 12
   2381: 'PH426 5P OUT OF RANGE', class Tank Control Warnings, trigger "2062_Warning_Data_BTCS_WARNING_WORD_16" bit 13
   2382: 'PH425 5S OUT OF RANGE', class Tank Control Warnings, trigger "2062_Warning_Data_BTCS_WARNING_WORD_16" bit 14
   2383: 'PH426 6P OUT OF RANGE', class Tank Control Warnings, trigger "2062_Warning_Data_BTCS_WARNING_WORD_16" bit 15
   2384: '', class Tank Control Warnings, trigger "2062_Warning_Data_BTCS_WARNING_WORD_17" bit 0
   2385: '', class Tank Control Warnings, trigger "2062_Warning_Data_BTCS_WARNING_WORD_17" bit 1
   2386: '', class Tank Control Warnings, trigger "2062_Warning_Data_BTCS_WARNING_WORD_17" bit 2
   2387: '', class Tank Control Warnings, trigger "2062_Warning_Data_BTCS_WARNING_WORD_17" bit 3
   2388: '', class Tank Control Warnings, trigger "2062_Warning_Data_BTCS_WARNING_WORD_17" bit 4
   2389: '', class Tank Control Warnings, trigger "2062_Warning_Data_BTCS_WARNING_WORD_17" bit 5
   2390: '', class Tank Control Warnings, trigger "2062_Warning_Data_BTCS_WARNING_WORD_17" bit 6
   2391: '', class Tank Control Warnings, trigger "2062_Warning_Data_BTCS_WARNING_WORD_17" bit 7
   2392: 'DO427 3S OUT OF RANGE', class Tank Control Warnings, trigger "2062_Warning_Data_BTCS_WARNING_WORD_17" bit 8
   2393: 'DO428 4P OUT OF RANGE', class Tank Control Warnings, trigger "2062_Warning_Data_BTCS_WARNING_WORD_17" bit 9
   2394: 'DO427 4S OUT OF RANGE', class Tank Control Warnings, trigger "2062_Warning_Data_BTCS_WARNING_WORD_17" bit 10
   2395: 'DO428 5P OUT OF RANGE', class Tank Control Warnings, trigger "2062_Warning_Data_BTCS_WARNING_WORD_17" bit 11
   2396: 'DO427 5S OUT OF RANGE', class Tank Control Warnings, trigger "2062_Warning_Data_BTCS_WARNING_WORD_17" bit 12
   2397: 'DO428 6P OUT OF RANGE', class Tank Control Warnings, trigger "2062_Warning_Data_BTCS_WARNING_WORD_17" bit 13
   2398: 'DO427 6S OUT OF RANGE', class Tank Control Warnings, trigger "2062_Warning_Data_BTCS_WARNING_WORD_17" bit 14
   2399: 'DO428 APT OUT OF RANGE', class Tank Control Warnings, trigger "2062_Warning_Data_BTCS_WARNING_WORD_17" bit 15

graphic list "Pump": 1 'Pump0'; 2 'Pump1'; 3 'Pump2'

graphic list "Pump Ani": 1 'Pumpd'; 0 'Pump0'; 1 'Pump1'; 2 'Pump2'; 5 'Pumpd'

graphic list "IA Compressor": 0 'IA Compressor 00'; 1 'IA Compressor 01'; 2 'IA Compressor 02_1'; 3 'IA Compressor 0_1'

graphic list "Tank Process Stage": 0 'Graphic_186'; 1 'Graphic_187'; 2 'Graphic_188'; 3 'Graphic_189'; 4 'Graphic_190'; 5 'Graphic_191'; 6 'Graphic_192'; 7 'Graphic_186'; 7 'Graphic_216'

graphic list "Water Level Override": 0 'Graphic_217'; 1 'Graphic_218'; 2 'Graphic_217'

graphic list "GCU": 0 'Graphic_150'; 1 'Graphic_150'

graphic list "IGGS": 0 'Graphic_3'; 1 'Graphic_140'

graphic list "Process time Banner": 2..5 'Graphic_193'; 1 'Pre Dwell'; 2 'Graphic_193'

graphic list "New IA Compressor": 0 'Graphic_249'; 1 'Graphic_250'; 2 'Graphic_249'; 3 'Graphic_250'

graphic list "Tank Process Stage_II": 0 'INITIAL STATE'; 1 'Pre Dwell'; 2 'De-Oxygenation'; 3 'Graphic_189'; 4 'Graphic_190'; 5 'Graphic_191'; 6 'Graphic_192'; 7 'Graphic_186'

screen "Main Index" 480x228, template "Template_1"
   on GenerateScreen: "TitleUpdater"()
   GraphicView "Graphic view_1" at 117,4 size 244x221; Picture "Graphic_115"
   Button "HmiScreenItemData_2" at 101,48 size 85x40; TextOn 'IGG Plant'; TextOff 'IGGS Plant'
      on Release: ActivateScreen("IGGS Plant", 0)
   Button "HmiScreenItemData_19" at 292,49 size 85x40; TextOn 'IGG Plant'; TextOff 'Alarms'
      on Release: ActivateScreen("Alarms", 0)
   Button "HmiScreenItemData_1" at 0,1 size 75x40; TextOn 'Back'; TextOff 'Home'
      on Release: ActivateScreen("Home", 0)
   Button "HmiScreenItemData_6" at 292,168 size 85x40; TextOn 'IGG Plant'; TextOff 'System Info'
      on Press: function_efd93a16("Info", 0, 0, -1, 3, 1)
   Button "HmiScreenItemData_3" at 197,48 size 85x40; TextOn 'IGG Plant'; TextOff 'BWTS'
      on Release: ActivateScreen("BWTS", 0)
   Button "HmiScreenItemData_11" at 197,107 size 85x40; TextOn 'IGG Plant'; TextOff 'GCU Plant'
      on Release: ActivateScreen("GCU Plant", 0)
   Button "HmiScreenItemData_10" at 197,168 size 85x40; TextOn 'IGG Plant'; TextOff 'PGC System'
      on Release: ActivateScreen("PGC", 0)
   Button "HmiScreenItemData_4" at 101,107 size 85x40; TextOn 'IGG Plant'; TextOff 'Air System'
      on Release: ActivateScreen("Air System", 0)
   Button "HmiScreenItemData_7" at 99,168 size 85x40; TextOn 'IGG Plant'; TextOff 'Fuel System'
      on Release: ActivateScreen("Fuel System", 0)
   Button "HmiScreenItemData_8" at 292,107 size 85x40; TextOn 'IGG Plant'; TextOff 'Cooling System'
      on Release: ActivateScreen("Cooling System", 0)

screen "Home" 480x228, template "Template_1"
   on GenerateScreen: "TitleUpdater"()
   Button "HmiScreenItemData" at 17,12 size 444x204; TextOn 'Main Index'; TextOff 'Text'
      on Release: ActivateScreen("Main Index", 0)
   GraphicView "Graphic view_2" at 19,14 size 100x200; Picture "Graphic_137"
   GraphicView "Graphic view_1" at 118,96 size 241x108; Picture "Graphic_185"
   TextField "HmiScreenItemData_3" at 76,57 size 326x26; Text 'Ballast Water Treatment System'
   TextField "HmiScreenItemData_4" at 53,27 size 371x29; Text 'Welcome to Coldharbour Marine'
   Circle "Circle_45" at 371,188 size 26x26
      Visibility <- "TRUE"
      Appearance <- "BRIGE HMI HEART BEAT"
   Circle "Circle_46" at 402,188 size 26x26
      Visibility <- "TRUE"
      Appearance <- "IGG PLC HEART BEAT"
   Button "Button_1" at 1,2 size 478x225; TextOff 'Text'
      on Release: ActivateScreen("Main Index", 0)
   Button "Button_2" at 436,194 size 44x34; TextOff 'Text'; PictureOff "Graphic_286"
      on Release: StopRuntime(0)

screen "GCU Plant" 480x228, template "Template_1"
   on GenerateScreen: "TitleUpdater"()
   Button "HmiScreenItemData_6" at 0,0 size 126x30; TextOn 'I&A Compressor Ok'; TextOff 'Previous Screen'
      on Release: function_efd93a16()
   GraphicView "Graphic view_1" at 138,24 size 127x184; Picture "Graphic_150"
   GraphicView "Graphic view_85" at 108,80 size 31x32; Picture "Graphic_178"
   GraphicView "Graphic view_87" at 107,102 size 18x56; Picture "Graphic_147"
   GraphicView "Graphic view_86" at 93,150 size 32x32; Picture "Graphic_159"
   Circle "Circle_1" at 109,167 size 6x6
      Visibility <- "10_DI_DATA_E_400_RUN"
      DiagonalMovement <- "E-400 Animation_DB_Animation"
   Circle "Circle_2" at 112,88 size 6x6
      Visibility <- "10_DI_DATA_E_400_RUN"
      VerticalMovement <- "E-400 Animation_DB_Animation"
   GraphicView "Graphic view_11" at 204,204 size 12x23; Picture "Graphic_152"
   Circle "Circle_31" at 155,85 size 6x6
      Visibility <- "10_DI_DATA_E_400_RUN"
      HorizontalMovement <- "E-400 Animation_DB_Animation"
   Circle "Circle_32" at 155,129 size 6x6
      Visibility <- "10_DI_DATA_E_400_RUN"
      DiagonalMovement <- "E-400 Animation_DB_Animation"
   Circle "Circle_33" at 179,152 size 6x6
      Visibility <- "10_DI_DATA_E_400_RUN"
      DiagonalMovement <- "E-400 Animation_DB_Animation"
   Circle "Circle_38" at 192,46 size 6x6
      Visibility <- "10_DI_DATA_E_400_RUN"
      DiagonalMovement <- "E-400 Animation_DB_Animation"
   Circle "Circle_39" at 223,52 size 6x6
      Visibility <- "10_DI_DATA_E_400_RUN"
      DiagonalMovement <- "E-400 Animation_DB_Animation"
   Circle "Circle_40" at 211,42 size 6x6
      Visibility <- "10_DI_DATA_E_400_RUN"
      DiagonalMovement <- "E-400 Animation_DB_Animation"
   Circle "Circle_41" at 224,36 size 6x6
      Visibility <- "10_DI_DATA_E_400_RUN"
      DiagonalMovement <- "E-400 Animation_DB_Animation"
   GraphicView "Graphic view_54" at 292,4 size 14x32; Picture "Graphic_147"
   GraphicView "Graphic view_2" at 258,34 size 182x14; Picture "Graphic_151"
   Circle "Circle_23" at 306,37 size 6x6
      Visibility <- "10_DI_DATA_E_400_RUN"
      HorizontalMovement <- "E-400 Animation_DB_Animation"
   Circle "Circle_24" at 318,40 size 6x6
      Visibility <- "10_DI_DATA_E_400_RUN"
      HorizontalMovement <- "E-400 Animation_DB_Animation"
   TextField "Text field_1" at 410,49 size 62x20; Text 'To Deck'
   TextField "Text field_2" at 0,155 size 45x36; Text 'From PGC'
   TextField "Text field_3" at 306,1 size 62x20; Text 'To Vent'
   GraphicView "Graphic view_3" at 50,163 size 34x19; Picture "Graphic_245"
   GraphicView "Graphic view_4" at 440,31 size 34x19; Picture "Graphic_245"
   Bar "Bar_1" at 186,61 size 48x135; Unit  %; MinimumValue 0; MaximumValue 100
      ProcessValue <- "12_AI_Data_LIT_304_SCALED"
   Button "HmiScreenItemData_2" at 399,4 size 80x25; TextOn 'IGG Plant'; TextOff 'BWTS'
      on Release: ActivateScreen("BWTS", 0)
   Button "HmiScreenItemData_3" at 0,196 size 80x25; TextOn 'IGG Plant'; TextOff 'PGC'
      on Release: ActivateScreen("PGC", 0)
   Circle "Circle_34" at 194,151 size 6x6
      DiagonalMovement <- "E-400 Animation_DB_Animation"
      Visibility <- "10_DI_DATA_E_400_RUN"
   Circle "Circle_37" at 198,129 size 6x6
      DiagonalMovement <- "E-400 Animation_DB_Animation"
      Visibility <- "10_DI_DATA_E_400_RUN"
   Circle "Circle_36" at 223,129 size 6x6
      DiagonalMovement <- "E-400 Animation_DB_Animation"
      Visibility <- "10_DI_DATA_E_400_RUN"
   Circle "Circle_35" at 205,175 size 6x6
      DiagonalMovement <- "E-400 Animation_DB_Animation"
      Visibility <- "10_DI_DATA_E_400_RUN"
   Button "HmiScreenItemData_1" at 1,34 size 84x30; TextOn 'I&A Compressor Ok'; TextOff 'Main Index'
      on Release: ActivateScreen("Main Index", 0)

screen "IGGS Plant" 480x228, template "Template_1"
   on GenerateScreen: "TitleUpdater"()
   Group "Group" at 8,32 size 343x170; Picture "Graphic_69"
   GraphicView "Graphic view_68" at 294,161 size 9x6; Picture "Graphic_107"
   GraphicView "Graphic view_36" at 303,36 size 18x23; Picture "Graphic_108"
   GraphicView "Graphic view_60" at 308,53 size 10x19; Picture "Graphic_17"
   GraphicView "Graphic view_4" at 260,36 size 16x23; Picture "Graphic_108"
   GraphicView "Graphic view_83" at 178,88 size 95x82; Picture "Graphic_130"
      Visibility <- "Flame"
   GraphicView "Graphic view_85" at 189,103 size 67x46; Picture "Graphic_132"
      Visibility <- "103_Main_Burner_DB_DN_OK"
   GraphicView "Graphic view_82" at 180,93 size 89x69; Picture "Graphic_130"
      Visibility <- "103_Main_Burner_DB_RUNNING"
   TextField "Text field_69" at 358,65 size 54x17; Text 'Oxygen'
   IOField "I/O field_22" at 413,64 size 62x20; FormatPattern 99.9; Unit  %
      ProcessValue <- "O2 Analyser Content Scaled"
   TextField "Text field_71" at 358,92 size 61x17; Text 'Setpoint'
   TextField "Text field_72" at 358,119 size 35x17; Text 'Soot'
   IOField "I/O field_24" at 413,118 size 62x20; FormatPattern 999; Unit  %
      ProcessValue <- "IG Soot Content Scaled"
   IOField "I/O field_25" at 413,145 size 62x20; FormatPattern 99; Unit  °C
      ProcessValue <- "Inert Gas Temp Scaled"
   TextField "Text field_73" at 358,145 size 45x17; Text 'Temp.'
   IOField "I/O field_26" at 413,173 size 62x20; FormatPattern 999; Unit  mBar
      ProcessValue <- "Inert Gas Pressure (PIT402) Scaled"
   TextField "Text field_74" at 358,172 size 45x17; Text 'Press.'
   IOField "I/O field_17" at 193,117 size 36x14; FormatPattern 999; Unit %
      ProcessValue <- "Flame Signal Scaled"
   Line "Line_4" at 190,102 size 1x7
      Visibility <- "Igniter Control"
   GraphicView "Graphic view_84" at 184,100 size 14x26; Picture "Graphic_129"
      Visibility <- "Pilot Flame"
   IOField "I/O field_23" at 413,91 size 62x20; Authorization "User administration"; FormatPattern 99.9; Unit  %
      ProcessValue <- "HMI Data_O2 Setpoint"
   TextField "Text field_70" at 357,40 size 121x18; Text 'Inert Gas Profile'
   Button "HmiScreenItemData_13" at 139,198 size 197x25; TextOn 'Back'; TextOff 'Cooling System'
      on Release: ActivateScreen("Cooling System", 0)
   Button "HmiScreenItemData_18" at 139,198 size 197x25; TextOn 'Back'; TextOff 'Cooling System'
      on Release: ActivateScreen("Cooling System", 0)
      Visibility <- "CSW Pump Control"
   Button "Button_2" at 1,61 size 115x25; TextOff 'Compressed Air'
      on Release: ActivateScreen("Air System", 0)
   Button "Button_5" at 1,98 size 115x25; TextOff 'Fuel System'
      on Release: ActivateScreen("Fuel System", 0)
   Button "Button_6" at 1,133 size 115x25; TextOff 'Combustion Air'
      on Release: ActivateScreen("CA Blower", 0)
   Button "Button_1" at 1,61 size 115x25; TextOff 'Compressed Air'
      on Release: ActivateScreen("Air System", 0)
      Visibility <- "Data_From BC PLC_Data_IA Compressor Running"
   Button "Button_3" at 1,98 size 115x25; TextOff 'Fuel System'
      on Release: ActivateScreen("Fuel System", 0)
      Visibility <- "Data To IGG PLC_Data_Fuel Oil System Proved"
   Button "Button_4" at 1,133 size 115x25; TextOff 'Combustion Air'
      on Release: ActivateScreen("CA Blower", 0)
      Visibility <- "CA Blower Running"
   Button "HmiScreenItemData_2" at 353,1 size 126x30; TextOn 'I&A Compressor Ok'; TextOff 'Previous Screen'
      on Release: function_efd93a16()
   Button "HmiScreenItemData_19" at 0,169 size 85x40; TextOn 'IGG Plant'; TextOff 'Alarms'
      on Release: ActivateScreen("Alarms", 0)
   Group "Group_12" at 129,1 size 89x43
   Circle "Circle_73" at 187,115 size 2x2
      HorizontalMovement <- "CA Blower Animation"
      Visibility <- "CA Blower On"
   Button "HmiScreenItemData_1" at 1,1 size 84x30; TextOn 'I&A Compressor Ok'; TextOff 'Main Index'
      on Release: ActivateScreen("Main Index", 0)
   Circle "Circle_98" at 258,155 size 8x8
      DiagonalMovement <- "CSW_Animation_DB_Animation"
      Visibility <- "Jacket Cooling Water Flow Switch"
   Circle "Circle_99" at 279,147 size 8x8
      DiagonalMovement <- "CSW_Animation_DB_Animation"
      Visibility <- "Jacket Cooling Water Flow Switch"
   Circle "Circle_104" at 261,133 size 8x8
      DiagonalMovement <- "CSW_Animation_DB_Animation"
      Visibility <- "Jacket Cooling Water Flow Switch"
   Circle "Circle_105" at 271,117 size 8x8
      DiagonalMovement <- "CSW_Animation_DB_Animation"
      Visibility <- "Jacket Cooling Water Flow Switch"
   Circle "Circle_107" at 276,137 size 8x8
      DiagonalMovement <- "CSW_Animation_DB_Animation"
      Visibility <- "Jacket Cooling Water Flow Switch"
   Circle "Circle_94" at 265,88 size 6x6
      DiagonalMovement <- "CSW_Animation_DB_Animation"
      Visibility <- "Jacket Cooling Water Flow Switch"
   Circle "Circle_100" at 276,162 size 8x8
      DiagonalMovement <- "CSW_Animation_DB_Animation"
      Visibility <- "Jacket Cooling Water Flow Switch"
   GraphicView "Graphic view_20" at 13,32 size 338x170; Picture "Graphic_69"
   Button "HmiScreenItemData_3" at 129,1 size 89x43; TextOn 'Back'; TextOff 'Burner Off'
      Visibility <- "103_Main_Burner_DB_Status"
   Button "HmiScreenItemData_4" at 129,1 size 89x43; TextOn 'Back'; TextOff 'Start Burner'
      Visibility <- "103_Main_Burner_DB_Status"
   Button "HmiScreenItemData_5" at 129,1 size 89x43; TextOn 'Back'; TextOff 'Burner On'
      Visibility <- "103_Main_Burner_DB_Status"
   Button "HmiScreenItemData_7" at 129,1 size 89x43; TextOn 'Back'; TextOff 'Burner Stopped'
      Visibility <- "103_Main_Burner_DB_Status"